// TIA Portal project "SSA-3GHz_V18" (V18) (continued)
       "SLI_gDB_T_CONFIG_PLC".configData.deviceIP.InterfaceAddress.ADDR[1] := 192;
       "SLI_gDB_T_CONFIG_PLC".configData.deviceIP.InterfaceAddress.ADDR[2] := 168;
       "SLI_gDB_T_CONFIG_PLC".configData.deviceIP.InterfaceAddress.ADDR[3] := 1;
       "SLI_gDB_T_CONFIG_PLC".configData.deviceIP.InterfaceAddress.ADDR[4] := 234;
       "SLI_gDB_T_CONFIG_PLC".configData.deviceIP.SubnetMask.ADDR[1] := 255;
       "SLI_gDB_T_CONFIG_PLC".configData.deviceIP.SubnetMask.ADDR[2] := 255;
       "SLI_gDB_T_CONFIG_PLC".configData.deviceIP.SubnetMask.ADDR[3] := 255;
       "SLI_gDB_T_CONFIG_PLC".configData.deviceIP.SubnetMask.ADDR[4] := 0;
       "SLI_gDB_T_CONFIG_PLC".configData.deviceIP.DefaultRouter.ADDR[1] := 192;
       "SLI_gDB_T_CONFIG_PLC".configData.deviceIP.DefaultRouter.ADDR[2] := 168;
       "SLI_gDB_T_CONFIG_PLC".configData.deviceIP.DefaultRouter.ADDR[3] := 1;
       "SLI_gDB_T_CONFIG_PLC".configData.deviceIP.DefaultRouter.ADDR[4] := 1;
   END_IF;
END_REGION

REGION Network 2: Set "start" to TRUE to configure the PROFINET interface.
   #_w1 := "tmp_setIP" AND NOT "Pulse_mem";   // rising edge of "tmp_setIP"
   "Pulse_mem" := "tmp_setIP";
   #_w2 := #_w1 OR "Set_IP_PArameters" OR "FirstScan" OR "RestoreFactorySettings";
   IF #_w2 THEN
       "SLI_gDB_T_CONFIG_PLC".T_CONFIG.start := TRUE;
       "Set_IP_PArameters" := FALSE;
   END_IF;
   "IEC_Timer_0_DB".TP(IN := #_w2, PT := t#5s);
   "ModbusData".serverData.disconnect := "IEC_Timer_0_DB".Q;
END_REGION

REGION Network 3: Set "start" to TRUE to configure the PROFINET interface.
   // NOTE! Before using the example:
   // 
   // Condition:
   // 1) Open the device view of the CPU "> Properties > PROFINET interface > Ethernet addresses > PROFINET". 
   // 2) To set the device name: Activate the following options: 
   // - "IP address is set directly at the device". 
   // - "PROFINET device name is set directly at the device".
   // 
   // Regarding parameter INTERFACE ("hwid"):
   // - Change the value of "hwid" according to the identification number of the PROFINET interface of your local device (CPU). (Open "PLC tags > Show all tags > System constants. Look for a name like "<Local~PROFINET_interface_1>" with a Data type "Hw_Interface". The cell "value" contains the hwid.)
   // 
   // Info:
   // In the "header" (IF_CONF_HEADER):
   // - SubfieldCount = 2: Indicates that two additional structures ("deviceIP" and "deviceName") are used below.
   // 
   // In the structure "deviceIP" (system data type IF_CONF_v4):
   // - Lenght = 18: Information on overall length of the structure (12 bytes for the device IP + 6 bytes for the parameters Id, Length and Mode)
   // - Mode = 1: Permanent change of the device IP.
   // - InterfaceAddress, SubnetMask, DefaultRouter: IP connection data.
   // 
   // In the structure "deviceName" (system data type IF_CONF_NOS):
   // - Lenght = 11: Information on overall length of the structure (5 bytes for the device name "myplc" + 6 bytes for the parameters Id, Length and Mode)
   // - Mode = 1: Permanent change of the device name in "myplc".
   // - NOS[1] ... NOS[5]: Device name (1 character / byte)
   // 
   // Note: Instead of an absolute length, you can use the default start value (Lenght = 0) for a dynamic length.
   // ENO of a box is taken as its EN; it also drops when the box reports an error
   "T_CONFIG_DB_PLC"(Req := "SLI_gDB_T_CONFIG_PLC".T_CONFIG.start,   // T_CONFIG
                     Interface := "SLI_gDB_T_CONFIG_PLC".T_CONFIG.hwid,
                     Conf_Data := "SLI_gDB_T_CONFIG_PLC".configData,
                     Done => #done_PLC,
                     Busy => "SLI_gDB_T_CONFIG_PLC".T_CONFIG.busy,
                     Error => "SLI_gDB_T_CONFIG_PLC".T_CONFIG.error,
                     Status => "SLI_gDB_T_CONFIG_PLC".T_CONFIG.status,
                     Err_Loc => #errorLocation_PLC);
   IF #done_PLC THEN "SLI_gDB_T_CONFIG_PLC".T_CONFIG.done := TRUE; END_IF;
END_REGION

REGION Network 4: INFO: Saves the value of "T_CONFIG.status" in case of an error of T_CONFIG in "T_CONFIG.memErrStat".
   RUNG wire#powerrail
      Contact( "SLI_gDB_T_CONFIG_PLC".T_CONFIG.error )
      Move(in := "SLI_gDB_T_CONFIG_PLC".T_CONFIG.status, out1 => "SLI_gDB_T_CONFIG_PLC".T_CONFIG.memErrStat)
      Move(in := #errorLocation_PLC, out1 => "SLI_gDB_T_CONFIG_PLC".T_CONFIG.errorLocation)
      R_Coil( "SLI_gDB_T_CONFIG_PLC".T_CONFIG.start )
   END_RUNG
   // the same network as SCL:
   IF "SLI_gDB_T_CONFIG_PLC".T_CONFIG.error THEN
       "SLI_gDB_T_CONFIG_PLC".T_CONFIG.memErrStat := "SLI_gDB_T_CONFIG_PLC".T_CONFIG.status;
       "SLI_gDB_T_CONFIG_PLC".T_CONFIG.errorLocation := #errorLocation_PLC;
       "SLI_gDB_T_CONFIG_PLC".T_CONFIG.start := FALSE;
   END_IF;
END_REGION

REGION Network 5: INFO: If T_CONFIG is done, "start" will be reset.
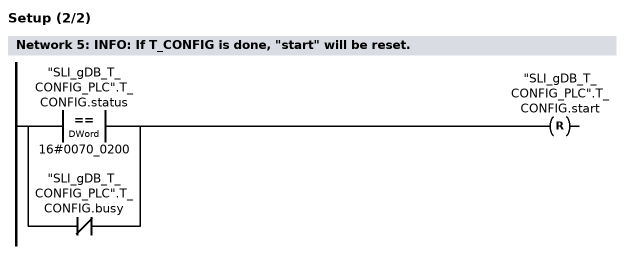
   RUNG wire#powerrail
      { S7_Templates := "SrcType := DWord" } EQ_Contact(in1 := "SLI_gDB_T_CONFIG_PLC".T_CONFIG.status, in2 := 16#0070_0200)
      wire#w1
      R_Coil( "SLI_gDB_T_CONFIG_PLC".T_CONFIG.start )
   END_RUNG
   RUNG wire#powerrail
      I_Contact( "SLI_gDB_T_CONFIG_PLC".T_CONFIG.busy )
   END_RUNG wire#w1
   // the same network as SCL:
   IF ("SLI_gDB_T_CONFIG_PLC".T_CONFIG.status = 16#0070_0200) OR NOT "SLI_gDB_T_CONFIG_PLC".T_CONFIG.busy THEN
       "SLI_gDB_T_CONFIG_PLC".T_CONFIG.start := FALSE;
   END_IF;
END_REGION
END_FUNCTION

FUNCTION "ProcessDI" : Void   // FC400, LAD
{ S7_Optimized_Access := 'TRUE' }
VERSION : 0.1
BEGIN

REGION Network 1: DutyCycOK
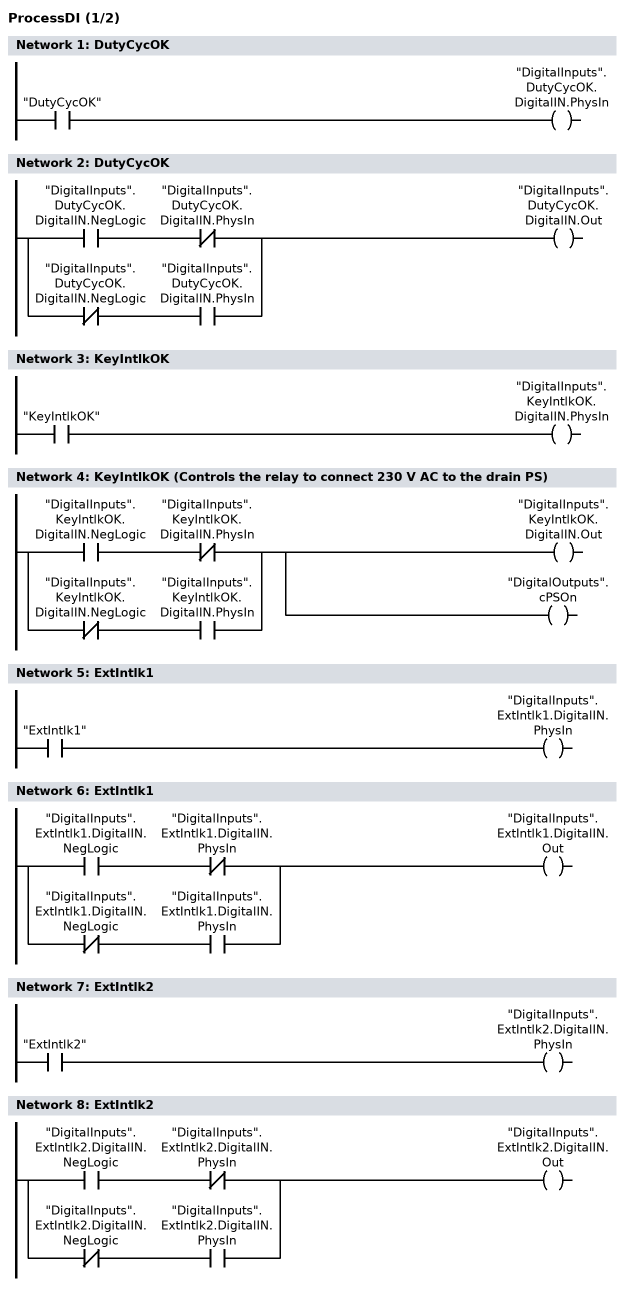
   RUNG wire#powerrail
      Contact( "DutyCycOK" )
      Coil( "DigitalInputs".DutyCycOK.DigitalIN.PhysIn )
   END_RUNG
   // the same network as SCL:
   "DigitalInputs".DutyCycOK.DigitalIN.PhysIn := "DutyCycOK";
END_REGION

REGION Network 2: DutyCycOK
   RUNG wire#powerrail
      Contact( "DigitalInputs".DutyCycOK.DigitalIN.NegLogic )
      I_Contact( "DigitalInputs".DutyCycOK.DigitalIN.PhysIn )
      wire#w1
      Coil( "DigitalInputs".DutyCycOK.DigitalIN.Out )
   END_RUNG
   RUNG wire#powerrail
      I_Contact( "DigitalInputs".DutyCycOK.DigitalIN.NegLogic )
      Contact( "DigitalInputs".DutyCycOK.DigitalIN.PhysIn )
   END_RUNG wire#w1
   // the same network as SCL:
   "DigitalInputs".DutyCycOK.DigitalIN.Out := ("DigitalInputs".DutyCycOK.DigitalIN.NegLogic AND NOT "DigitalInputs".DutyCycOK.DigitalIN.PhysIn) OR (NOT "DigitalInputs".DutyCycOK.DigitalIN.NegLogic AND "DigitalInputs".DutyCycOK.DigitalIN.PhysIn);
END_REGION

REGION Network 3: KeyIntlkOK
   RUNG wire#powerrail
      Contact( "KeyIntlkOK" )
      Coil( "DigitalInputs".KeyIntlkOK.DigitalIN.PhysIn )
   END_RUNG
   // the same network as SCL:
   "DigitalInputs".KeyIntlkOK.DigitalIN.PhysIn := "KeyIntlkOK";
END_REGION

REGION Network 4: KeyIntlkOK (Controls the relay to connect 230 V AC to the drain PS)
   RUNG wire#powerrail
      Contact( "DigitalInputs".KeyIntlkOK.DigitalIN.NegLogic )
      I_Contact( "DigitalInputs".KeyIntlkOK.DigitalIN.PhysIn )
      wire#w1
      Coil( "DigitalInputs".KeyIntlkOK.DigitalIN.Out )
   END_RUNG
   RUNG wire#powerrail
      I_Contact( "DigitalInputs".KeyIntlkOK.DigitalIN.NegLogic )
      Contact( "DigitalInputs".KeyIntlkOK.DigitalIN.PhysIn )
   END_RUNG wire#w1
   RUNG wire#w1
      Coil( "DigitalOutputs".cPSOn )
   END_RUNG
   // the same network as SCL:
   "DigitalInputs".KeyIntlkOK.DigitalIN.Out := ("DigitalInputs".KeyIntlkOK.DigitalIN.NegLogic AND NOT "DigitalInputs".KeyIntlkOK.DigitalIN.PhysIn) OR (NOT "DigitalInputs".KeyIntlkOK.DigitalIN.NegLogic AND "DigitalInputs".KeyIntlkOK.DigitalIN.PhysIn);
   "DigitalOutputs".cPSOn := "DigitalInputs".KeyIntlkOK.DigitalIN.Out;
END_REGION

REGION Network 5: ExtIntlk1
   RUNG wire#powerrail
      Contact( "ExtIntlk1" )
      Coil( "DigitalInputs".ExtIntlk1.DigitalIN.PhysIn )
   END_RUNG
   // the same network as SCL:
   "DigitalInputs".ExtIntlk1.DigitalIN.PhysIn := "ExtIntlk1";
END_REGION

REGION Network 6: ExtIntlk1
   RUNG wire#powerrail
      Contact( "DigitalInputs".ExtIntlk1.DigitalIN.NegLogic )
      I_Contact( "DigitalInputs".ExtIntlk1.DigitalIN.PhysIn )
      wire#w1
      Coil( "DigitalInputs".ExtIntlk1.DigitalIN.Out )
   END_RUNG
   RUNG wire#powerrail
      I_Contact( "DigitalInputs".ExtIntlk1.DigitalIN.NegLogic )
      Contact( "DigitalInputs".ExtIntlk1.DigitalIN.PhysIn )
   END_RUNG wire#w1
   // the same network as SCL:
   "DigitalInputs".ExtIntlk1.DigitalIN.Out := ("DigitalInputs".ExtIntlk1.DigitalIN.NegLogic AND NOT "DigitalInputs".ExtIntlk1.DigitalIN.PhysIn) OR (NOT "DigitalInputs".ExtIntlk1.DigitalIN.NegLogic AND "DigitalInputs".ExtIntlk1.DigitalIN.PhysIn);
END_REGION

REGION Network 7: ExtIntlk2
   RUNG wire#powerrail
      Contact( "ExtIntlk2" )
      Coil( "DigitalInputs".ExtIntlk2.DigitalIN.PhysIn )
   END_RUNG
   // the same network as SCL:
   "DigitalInputs".ExtIntlk2.DigitalIN.PhysIn := "ExtIntlk2";
END_REGION

REGION Network 8: ExtIntlk2
   RUNG wire#powerrail
      Contact( "DigitalInputs".ExtIntlk2.DigitalIN.NegLogic )
      I_Contact( "DigitalInputs".ExtIntlk2.DigitalIN.PhysIn )
      wire#w1
      Coil( "DigitalInputs".ExtIntlk2.DigitalIN.Out )
   END_RUNG
   RUNG wire#powerrail
      I_Contact( "DigitalInputs".ExtIntlk2.DigitalIN.NegLogic )
      Contact( "DigitalInputs".ExtIntlk2.DigitalIN.PhysIn )
   END_RUNG wire#w1
   // the same network as SCL:
   "DigitalInputs".ExtIntlk2.DigitalIN.Out := ("DigitalInputs".ExtIntlk2.DigitalIN.NegLogic AND NOT "DigitalInputs".ExtIntlk2.DigitalIN.PhysIn) OR (NOT "DigitalInputs".ExtIntlk2.DigitalIN.NegLogic AND "DigitalInputs".ExtIntlk2.DigitalIN.PhysIn);
END_REGION

REGION Network 9: T1_OK
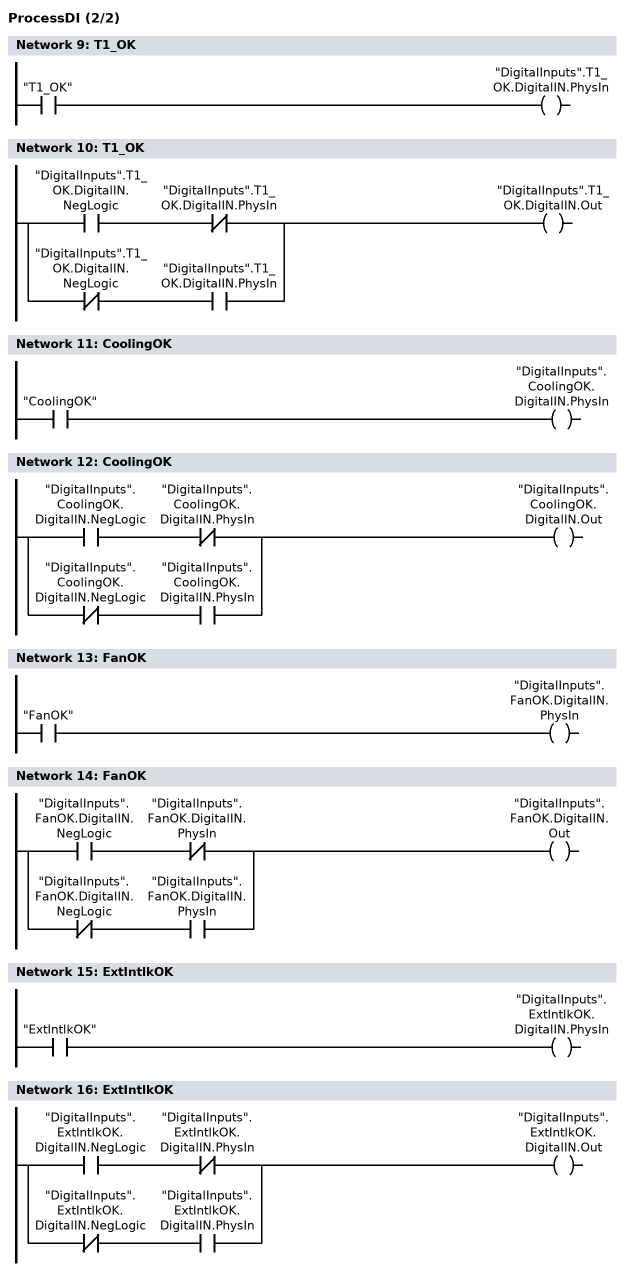
   RUNG wire#powerrail
      Contact( "T1_OK" )
      Coil( "DigitalInputs".T1_OK.DigitalIN.PhysIn )
   END_RUNG
   // the same network as SCL:
   "DigitalInputs".T1_OK.DigitalIN.PhysIn := "T1_OK";
END_REGION

REGION Network 10: T1_OK
   RUNG wire#powerrail
      Contact( "DigitalInputs".T1_OK.DigitalIN.NegLogic )
      I_Contact( "DigitalInputs".T1_OK.DigitalIN.PhysIn )
      wire#w1
      Coil( "DigitalInputs".T1_OK.DigitalIN.Out )
   END_RUNG
   RUNG wire#powerrail
      I_Contact( "DigitalInputs".T1_OK.DigitalIN.NegLogic )
      Contact( "DigitalInputs".T1_OK.DigitalIN.PhysIn )
   END_RUNG wire#w1
   // the same network as SCL:
   "DigitalInputs".T1_OK.DigitalIN.Out := ("DigitalInputs".T1_OK.DigitalIN.NegLogic AND NOT "DigitalInputs".T1_OK.DigitalIN.PhysIn) OR (NOT "DigitalInputs".T1_OK.DigitalIN.NegLogic AND "DigitalInputs".T1_OK.DigitalIN.PhysIn);
END_REGION

REGION Network 11: CoolingOK
   RUNG wire#powerrail
      Contact( "CoolingOK" )
      Coil( "DigitalInputs".CoolingOK.DigitalIN.PhysIn )
   END_RUNG
   // the same network as SCL:
   "DigitalInputs".CoolingOK.DigitalIN.PhysIn := "CoolingOK";
END_REGION

REGION Network 12: CoolingOK
   RUNG wire#powerrail
      Contact( "DigitalInputs".CoolingOK.DigitalIN.NegLogic )
      I_Contact( "DigitalInputs".CoolingOK.DigitalIN.PhysIn )
      wire#w1
      Coil( "DigitalInputs".CoolingOK.DigitalIN.Out )
   END_RUNG
   RUNG wire#powerrail
      I_Contact( "DigitalInputs".CoolingOK.DigitalIN.NegLogic )
      Contact( "DigitalInputs".CoolingOK.DigitalIN.PhysIn )
   END_RUNG wire#w1
   // the same network as SCL:
   "DigitalInputs".CoolingOK.DigitalIN.Out := ("DigitalInputs".CoolingOK.DigitalIN.NegLogic AND NOT "DigitalInputs".CoolingOK.DigitalIN.PhysIn) OR (NOT "DigitalInputs".CoolingOK.DigitalIN.NegLogic AND "DigitalInputs".CoolingOK.DigitalIN.PhysIn);
END_REGION

REGION Network 13: FanOK
   RUNG wire#powerrail
      Contact( "FanOK" )
      Coil( "DigitalInputs".FanOK.DigitalIN.PhysIn )
   END_RUNG
   // the same network as SCL:
   "DigitalInputs".FanOK.DigitalIN.PhysIn := "FanOK";
END_REGION

REGION Network 14: FanOK
   RUNG wire#powerrail
      Contact( "DigitalInputs".FanOK.DigitalIN.NegLogic )
      I_Contact( "DigitalInputs".FanOK.DigitalIN.PhysIn )
      wire#w1
      Coil( "DigitalInputs".FanOK.DigitalIN.Out )
   END_RUNG
   RUNG wire#powerrail
      I_Contact( "DigitalInputs".FanOK.DigitalIN.NegLogic )
      Contact( "DigitalInputs".FanOK.DigitalIN.PhysIn )
   END_RUNG wire#w1
   // the same network as SCL:
   "DigitalInputs".FanOK.DigitalIN.Out := ("DigitalInputs".FanOK.DigitalIN.NegLogic AND NOT "DigitalInputs".FanOK.DigitalIN.PhysIn) OR (NOT "DigitalInputs".FanOK.DigitalIN.NegLogic AND "DigitalInputs".FanOK.DigitalIN.PhysIn);
END_REGION

REGION Network 15: ExtIntlkOK
   RUNG wire#powerrail
      Contact( "ExtIntlkOK" )
      Coil( "DigitalInputs".ExtIntlkOK.DigitalIN.PhysIn )
   END_RUNG
   // the same network as SCL:
   "DigitalInputs".ExtIntlkOK.DigitalIN.PhysIn := "ExtIntlkOK";
END_REGION

REGION Network 16: ExtIntlkOK
   RUNG wire#powerrail
      Contact( "DigitalInputs".ExtIntlkOK.DigitalIN.NegLogic )
      I_Contact( "DigitalInputs".ExtIntlkOK.DigitalIN.PhysIn )
      wire#w1
      Coil( "DigitalInputs".ExtIntlkOK.DigitalIN.Out )
   END_RUNG
   RUNG wire#powerrail
      I_Contact( "DigitalInputs".ExtIntlkOK.DigitalIN.NegLogic )
      Contact( "DigitalInputs".ExtIntlkOK.DigitalIN.PhysIn )
   END_RUNG wire#w1
   // the same network as SCL:
   "DigitalInputs".ExtIntlkOK.DigitalIN.Out := ("DigitalInputs".ExtIntlkOK.DigitalIN.NegLogic AND NOT "DigitalInputs".ExtIntlkOK.DigitalIN.PhysIn) OR (NOT "DigitalInputs".ExtIntlkOK.DigitalIN.NegLogic AND "DigitalInputs".ExtIntlkOK.DigitalIN.PhysIn);
END_REGION
END_FUNCTION

FUNCTION "ProcessAI" : Void   // FC401, LAD
{ S7_Optimized_Access := 'TRUE' }
VERSION : 0.1
   VAR_TEMP
      tmpR1 : Real;
      tmpR : Real;
   END_VAR
BEGIN

REGION Network 1: U drain_RBK
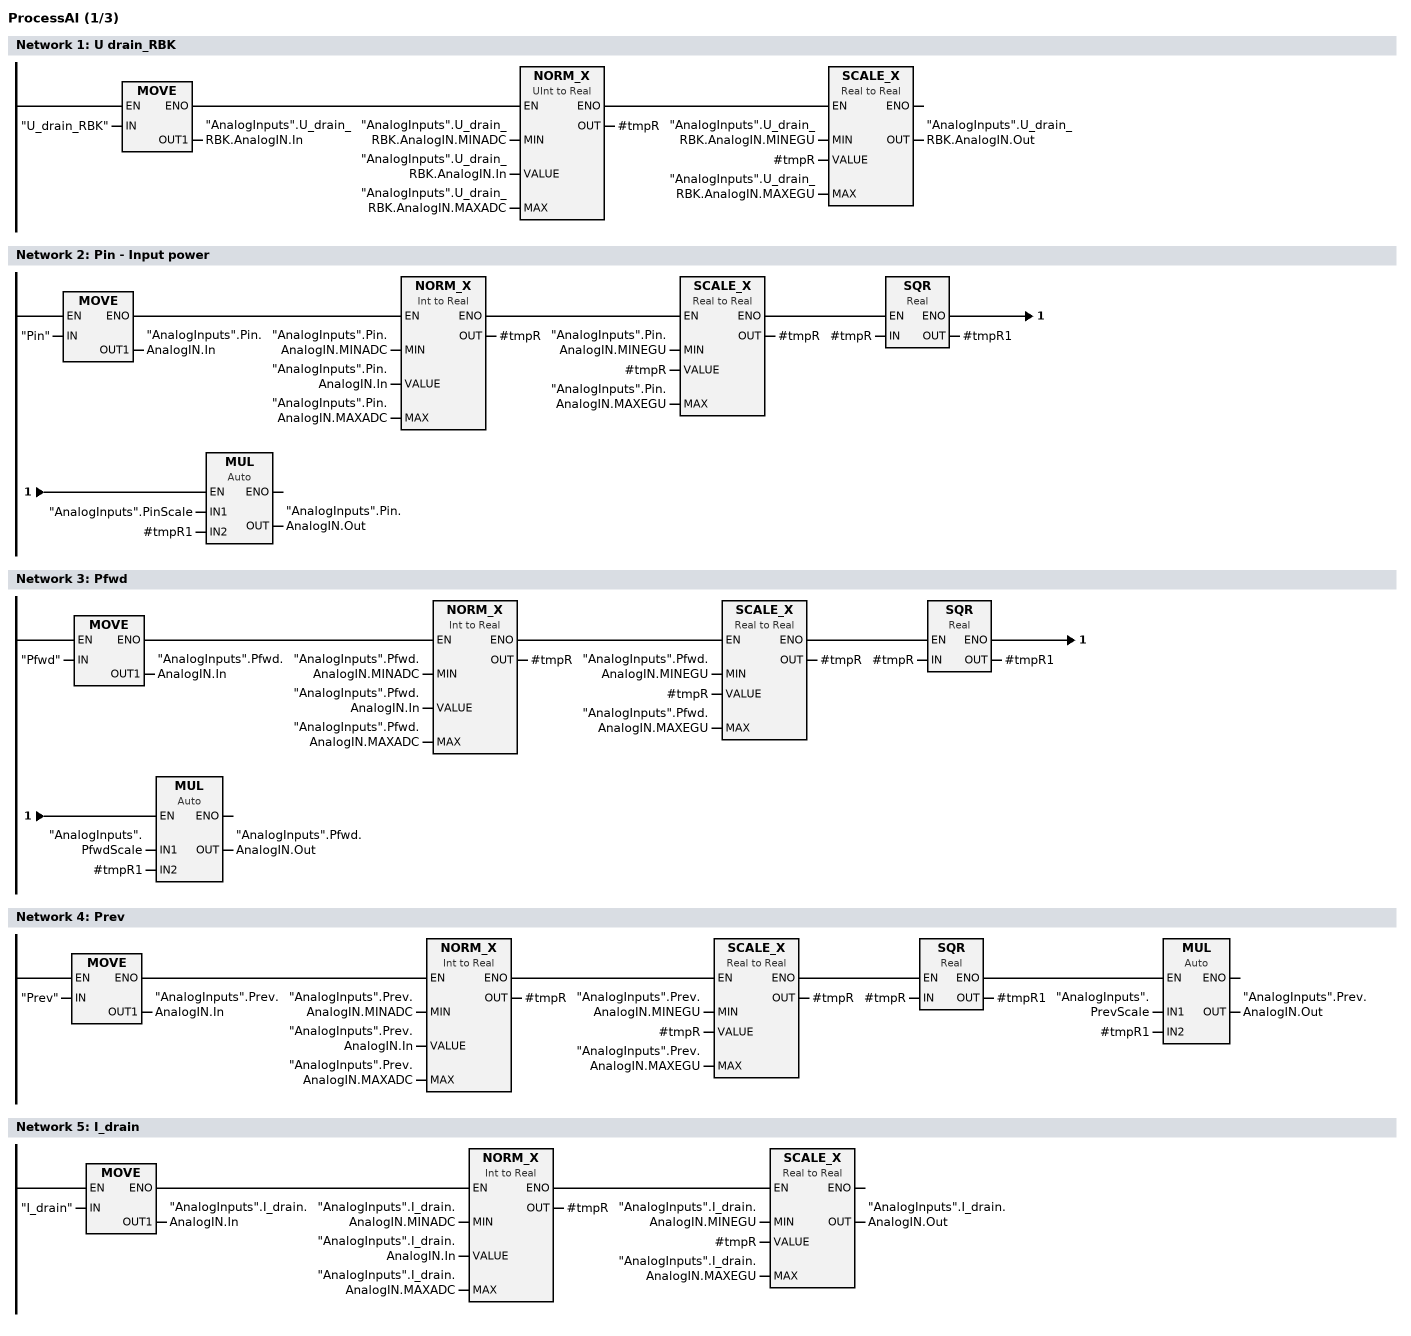
   RUNG wire#powerrail
      Move(in := "U_drain_RBK", out1 => "AnalogInputs".U_drain_RBK.AnalogIN.In)
      { S7_Templates := "[SrcType := UInt, DestType := Real]" } Normalize(min := "AnalogInputs".U_drain_RBK.AnalogIN.MINADC, value := "AnalogInputs".U_drain_RBK.AnalogIN.In, max := "AnalogInputs".U_drain_RBK.AnalogIN.MAXADC, out => #tmpR)
      { S7_Templates := "[SrcType := Real, DestType := Real]" } Scale(min := "AnalogInputs".U_drain_RBK.AnalogIN.MINEGU, value := #tmpR, max := "AnalogInputs".U_drain_RBK.AnalogIN.MAXEGU, out => "AnalogInputs".U_drain_RBK.AnalogIN.Out)
   END_RUNG
   // the same network as SCL:
   "AnalogInputs".U_drain_RBK.AnalogIN.In := "U_drain_RBK";
   #tmpR := NORM_X(MIN := "AnalogInputs".U_drain_RBK.AnalogIN.MINADC, VALUE := "AnalogInputs".U_drain_RBK.AnalogIN.In, MAX := "AnalogInputs".U_drain_RBK.AnalogIN.MAXADC);
   "AnalogInputs".U_drain_RBK.AnalogIN.Out := SCALE_X(MIN := "AnalogInputs".U_drain_RBK.AnalogIN.MINEGU, VALUE := #tmpR, MAX := "AnalogInputs".U_drain_RBK.AnalogIN.MAXEGU);
END_REGION

REGION Network 2: Pin - Input power
   "AnalogInputs".Pin.AnalogIN.In := "Pin";
   #tmpR := NORM_X(MIN := "AnalogInputs".Pin.AnalogIN.MINADC, VALUE := "AnalogInputs".Pin.AnalogIN.In, MAX := "AnalogInputs".Pin.AnalogIN.MAXADC);
   #tmpR := SCALE_X(MIN := "AnalogInputs".Pin.AnalogIN.MINEGU, VALUE := #tmpR, MAX := "AnalogInputs".Pin.AnalogIN.MAXEGU);
   #tmpR1 := SQR(#tmpR);
   "AnalogInputs".Pin.AnalogIN.Out := "AnalogInputs".PinScale * #tmpR1;
END_REGION

REGION Network 3: Pfwd
   "AnalogInputs".Pfwd.AnalogIN.In := "Pfwd";
   #tmpR := NORM_X(MIN := "AnalogInputs".Pfwd.AnalogIN.MINADC, VALUE := "AnalogInputs".Pfwd.AnalogIN.In, MAX := "AnalogInputs".Pfwd.AnalogIN.MAXADC);
   #tmpR := SCALE_X(MIN := "AnalogInputs".Pfwd.AnalogIN.MINEGU, VALUE := #tmpR, MAX := "AnalogInputs".Pfwd.AnalogIN.MAXEGU);
   #tmpR1 := SQR(#tmpR);
   "AnalogInputs".Pfwd.AnalogIN.Out := "AnalogInputs".PfwdScale * #tmpR1;
END_REGION

REGION Network 4: Prev
   "AnalogInputs".Prev.AnalogIN.In := "Prev";
   #tmpR := NORM_X(MIN := "AnalogInputs".Prev.AnalogIN.MINADC, VALUE := "AnalogInputs".Prev.AnalogIN.In, MAX := "AnalogInputs".Prev.AnalogIN.MAXADC);
   #tmpR := SCALE_X(MIN := "AnalogInputs".Prev.AnalogIN.MINEGU, VALUE := #tmpR, MAX := "AnalogInputs".Prev.AnalogIN.MAXEGU);
   #tmpR1 := SQR(#tmpR);
   "AnalogInputs".Prev.AnalogIN.Out := "AnalogInputs".PrevScale * #tmpR1;
END_REGION

REGION Network 5: I_drain
   RUNG wire#powerrail
      Move(in := "I_drain", out1 => "AnalogInputs".I_drain.AnalogIN.In)
      { S7_Templates := "[SrcType := Int, DestType := Real]" } Normalize(min := "AnalogInputs".I_drain.AnalogIN.MINADC, value := "AnalogInputs".I_drain.AnalogIN.In, max := "AnalogInputs".I_drain.AnalogIN.MAXADC, out => #tmpR)
      { S7_Templates := "[SrcType := Real, DestType := Real]" } Scale(min := "AnalogInputs".I_drain.AnalogIN.MINEGU, value := #tmpR, max := "AnalogInputs".I_drain.AnalogIN.MAXEGU, out => "AnalogInputs".I_drain.AnalogIN.Out)
   END_RUNG
   // the same network as SCL:
   "AnalogInputs".I_drain.AnalogIN.In := "I_drain";
   #tmpR := NORM_X(MIN := "AnalogInputs".I_drain.AnalogIN.MINADC, VALUE := "AnalogInputs".I_drain.AnalogIN.In, MAX := "AnalogInputs".I_drain.AnalogIN.MAXADC);
   "AnalogInputs".I_drain.AnalogIN.Out := SCALE_X(MIN := "AnalogInputs".I_drain.AnalogIN.MINEGU, VALUE := #tmpR, MAX := "AnalogInputs".I_drain.AnalogIN.MAXEGU);
END_REGION

REGION Network 6: ADC0ch1
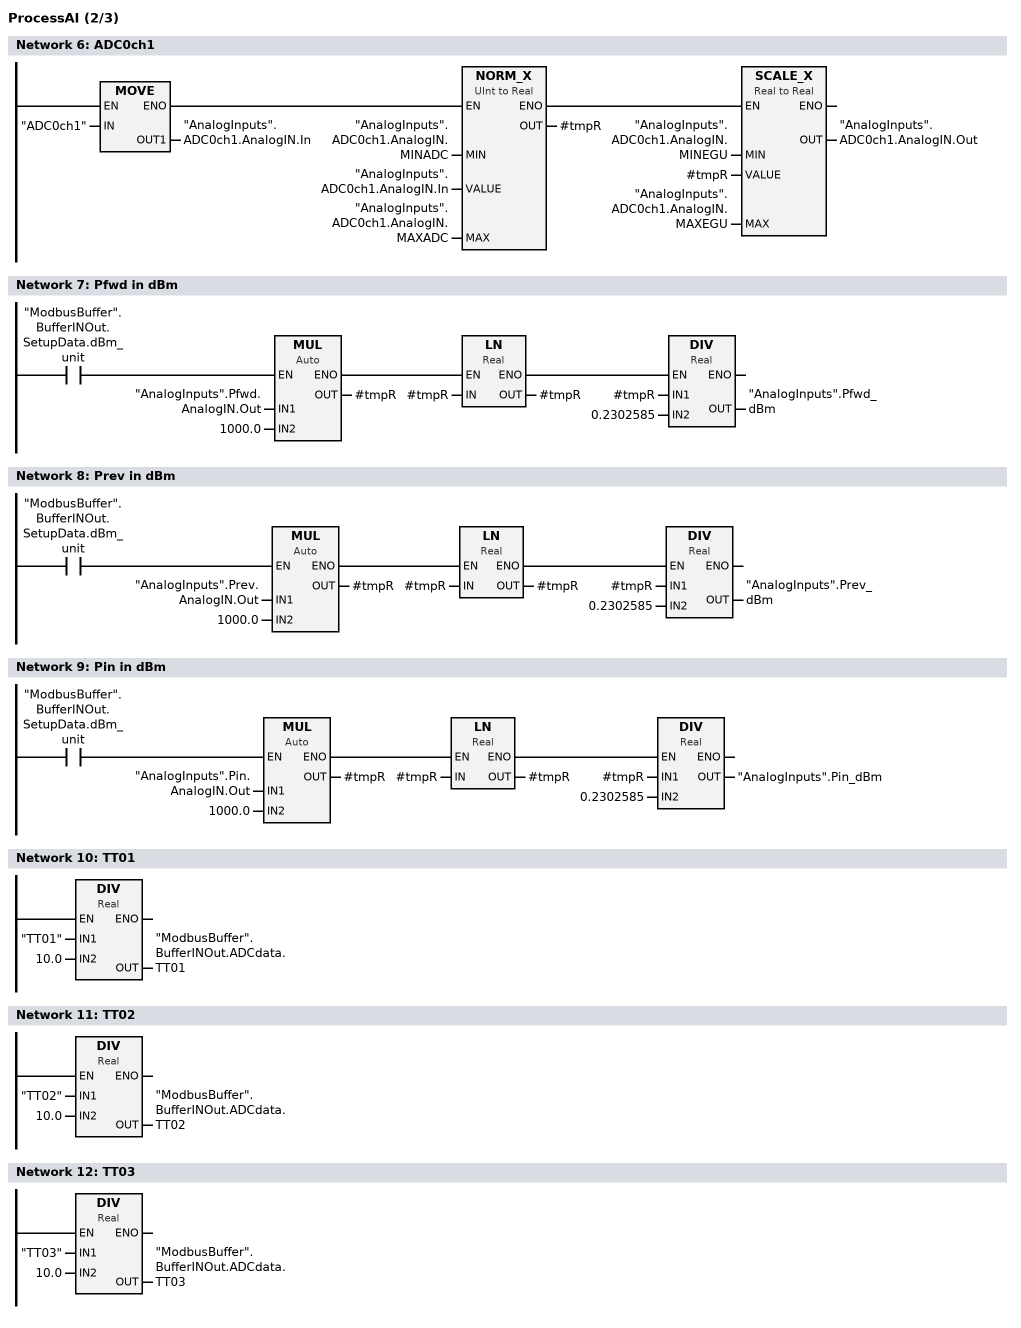
   RUNG wire#powerrail
      Move(in := "ADC0ch1", out1 => "AnalogInputs".ADC0ch1.AnalogIN.In)
      { S7_Templates := "[SrcType := UInt, DestType := Real]" } Normalize(min := "AnalogInputs".ADC0ch1.AnalogIN.MINADC, value := "AnalogInputs".ADC0ch1.AnalogIN.In, max := "AnalogInputs".ADC0ch1.AnalogIN.MAXADC, out => #tmpR)
      { S7_Templates := "[SrcType := Real, DestType := Real]" } Scale(min := "AnalogInputs".ADC0ch1.AnalogIN.MINEGU, value := #tmpR, max := "AnalogInputs".ADC0ch1.AnalogIN.MAXEGU, out => "AnalogInputs".ADC0ch1.AnalogIN.Out)
   END_RUNG
   // the same network as SCL:
   "AnalogInputs".ADC0ch1.AnalogIN.In := "ADC0ch1";
   #tmpR := NORM_X(MIN := "AnalogInputs".ADC0ch1.AnalogIN.MINADC, VALUE := "AnalogInputs".ADC0ch1.AnalogIN.In, MAX := "AnalogInputs".ADC0ch1.AnalogIN.MAXADC);
   "AnalogInputs".ADC0ch1.AnalogIN.Out := SCALE_X(MIN := "AnalogInputs".ADC0ch1.AnalogIN.MINEGU, VALUE := #tmpR, MAX := "AnalogInputs".ADC0ch1.AnalogIN.MAXEGU);
END_REGION

REGION Network 7: Pfwd in dBm
   IF "ModbusBuffer".BufferINOut.SetupData.dBm_unit THEN
       #tmpR := "AnalogInputs".Pfwd.AnalogIN.Out * 1000.0;
       #tmpR := LN(#tmpR);
       "AnalogInputs".Pfwd_dBm := #tmpR / 0.2302585;
   END_IF;
END_REGION

REGION Network 8: Prev in dBm
   IF "ModbusBuffer".BufferINOut.SetupData.dBm_unit THEN
       #tmpR := "AnalogInputs".Prev.AnalogIN.Out * 1000.0;
       #tmpR := LN(#tmpR);
       "AnalogInputs".Prev_dBm := #tmpR / 0.2302585;
   END_IF;
END_REGION

REGION Network 9: Pin in dBm
   IF "ModbusBuffer".BufferINOut.SetupData.dBm_unit THEN
       #tmpR := "AnalogInputs".Pin.AnalogIN.Out * 1000.0;
       #tmpR := LN(#tmpR);
       "AnalogInputs".Pin_dBm := #tmpR / 0.2302585;
   END_IF;
END_REGION

REGION Network 10: TT01
   RUNG wire#powerrail
      { S7_Templates := "SrcType := Real" } Div(in1 := "TT01", in2 := 10.0, out => "ModbusBuffer".BufferINOut.ADCdata.TT01)
   END_RUNG
   // the same network as SCL:
   "ModbusBuffer".BufferINOut.ADCdata.TT01 := "TT01" / 10.0;
END_REGION

REGION Network 11: TT02
   RUNG wire#powerrail
      { S7_Templates := "SrcType := Real" } Div(in1 := "TT02", in2 := 10.0, out => "ModbusBuffer".BufferINOut.ADCdata.TT02)
   END_RUNG
   // the same network as SCL:
   "ModbusBuffer".BufferINOut.ADCdata.TT02 := "TT02" / 10.0;
END_REGION

REGION Network 12: TT03
   RUNG wire#powerrail
      { S7_Templates := "SrcType := Real" } Div(in1 := "TT03", in2 := 10.0, out => "ModbusBuffer".BufferINOut.ADCdata.TT03)
   END_RUNG
   // the same network as SCL:
   "ModbusBuffer".BufferINOut.ADCdata.TT03 := "TT03" / 10.0;
END_REGION

REGION Network 13: TT04
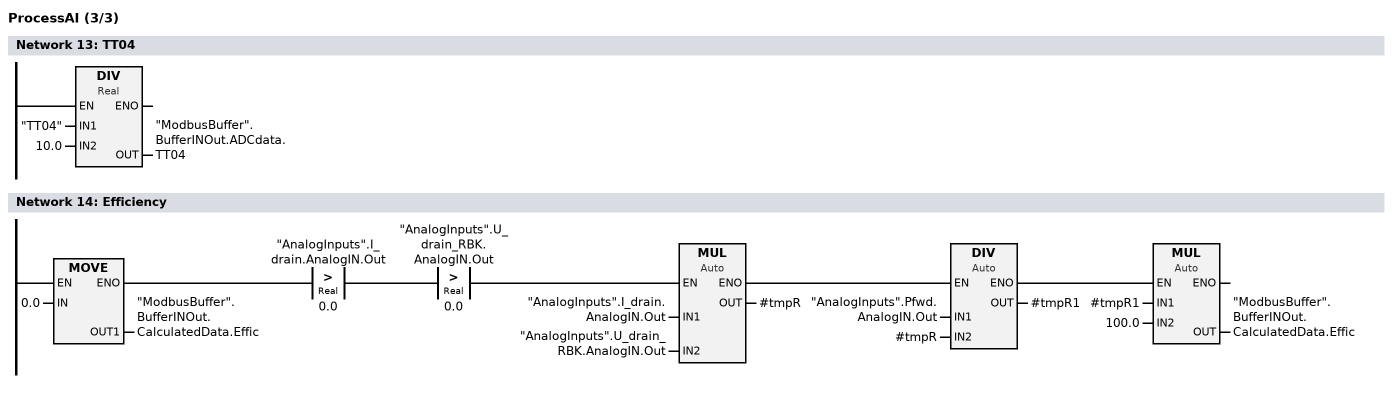
   RUNG wire#powerrail
      { S7_Templates := "SrcType := Real" } Div(in1 := "TT04", in2 := 10.0, out => "ModbusBuffer".BufferINOut.ADCdata.TT04)
   END_RUNG
   // the same network as SCL:
   "ModbusBuffer".BufferINOut.ADCdata.TT04 := "TT04" / 10.0;
END_REGION

REGION Network 14: Efficiency
   RUNG wire#powerrail
      Move(in := 0.0, out1 => "ModbusBuffer".BufferINOut.CalculatedData.Effic)
      { S7_Templates := "SrcType := Real" } GT_Contact(in1 := "AnalogInputs".I_drain.AnalogIN.Out, in2 := 0.0)
      { S7_Templates := "SrcType := Real" } GT_Contact(in1 := "AnalogInputs".U_drain_RBK.AnalogIN.Out, in2 := 0.0)
      Mul(in1 := "AnalogInputs".I_drain.AnalogIN.Out, in2 := "AnalogInputs".U_drain_RBK.AnalogIN.Out, out => #tmpR)
      Div(in1 := "AnalogInputs".Pfwd.AnalogIN.Out, in2 := #tmpR, out => #tmpR1)
      Mul(in1 := #tmpR1, in2 := 100.0, out => "ModbusBuffer".BufferINOut.CalculatedData.Effic)
   END_RUNG
   // the same network as SCL:
   "ModbusBuffer".BufferINOut.CalculatedData.Effic := 0.0;
   IF ("AnalogInputs".I_drain.AnalogIN.Out > 0.0) AND ("AnalogInputs".U_drain_RBK.AnalogIN.Out > 0.0) THEN
       #tmpR := "AnalogInputs".I_drain.AnalogIN.Out * "AnalogInputs".U_drain_RBK.AnalogIN.Out;
       #tmpR1 := "AnalogInputs".Pfwd.AnalogIN.Out / #tmpR;
       "ModbusBuffer".BufferINOut.CalculatedData.Effic := #tmpR1 * 100.0;
   END_IF;
END_REGION
END_FUNCTION

FUNCTION "ProcessAO" : Void   // FC402, LAD
{ S7_Optimized_Access := 'TRUE' }
VERSION : 0.1
   VAR_TEMP
      tmpR : Real;
   END_VAR
BEGIN

REGION Network 1: U drain
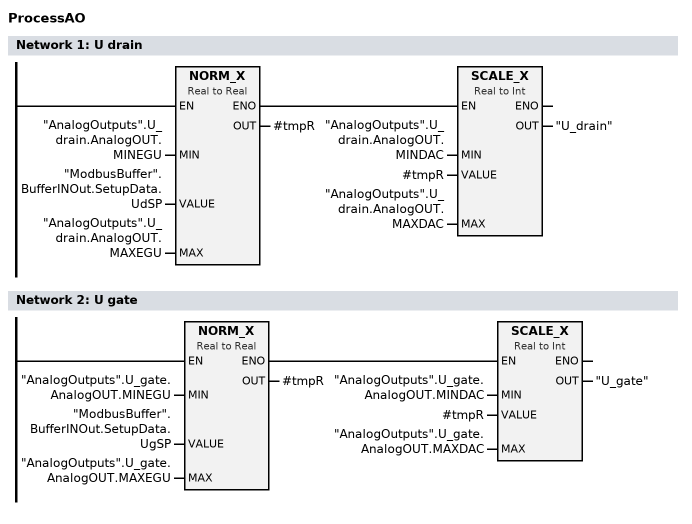
   RUNG wire#powerrail
      { S7_Templates := "[SrcType := Real, DestType := Real]" } Normalize(min := "AnalogOutputs".U_drain.AnalogOUT.MINEGU, value := "ModbusBuffer".BufferINOut.SetupData.UdSP, max := "AnalogOutputs".U_drain.AnalogOUT.MAXEGU, out => #tmpR)
      { S7_Templates := "[SrcType := Real, DestType := Int]" } Scale(min := "AnalogOutputs".U_drain.AnalogOUT.MINDAC, value := #tmpR, max := "AnalogOutputs".U_drain.AnalogOUT.MAXDAC, out => "U_drain")
   END_RUNG
   // the same network as SCL:
   #tmpR := NORM_X(MIN := "AnalogOutputs".U_drain.AnalogOUT.MINEGU, VALUE := "ModbusBuffer".BufferINOut.SetupData.UdSP, MAX := "AnalogOutputs".U_drain.AnalogOUT.MAXEGU);
   "U_drain" := SCALE_X(MIN := "AnalogOutputs".U_drain.AnalogOUT.MINDAC, VALUE := #tmpR, MAX := "AnalogOutputs".U_drain.AnalogOUT.MAXDAC);
END_REGION

REGION Network 2: U gate
   RUNG wire#powerrail
      { S7_Templates := "[SrcType := Real, DestType := Real]" } Normalize(min := "AnalogOutputs".U_gate.AnalogOUT.MINEGU, value := "ModbusBuffer".BufferINOut.SetupData.UgSP, max := "AnalogOutputs".U_gate.AnalogOUT.MAXEGU, out => #tmpR)
      { S7_Templates := "[SrcType := Real, DestType := Int]" } Scale(min := "AnalogOutputs".U_gate.AnalogOUT.MINDAC, value := #tmpR, max := "AnalogOutputs".U_gate.AnalogOUT.MAXDAC, out => "U_gate")
   END_RUNG
   // the same network as SCL:
   #tmpR := NORM_X(MIN := "AnalogOutputs".U_gate.AnalogOUT.MINEGU, VALUE := "ModbusBuffer".BufferINOut.SetupData.UgSP, MAX := "AnalogOutputs".U_gate.AnalogOUT.MAXEGU);
   "U_gate" := SCALE_X(MIN := "AnalogOutputs".U_gate.AnalogOUT.MINDAC, VALUE := #tmpR, MAX := "AnalogOutputs".U_gate.AnalogOUT.MAXDAC);
END_REGION
END_FUNCTION

FUNCTION "ProcessDO" : Void   // FC450, LAD
{ S7_Optimized_Access := 'TRUE' }
VERSION : 0.1
BEGIN

REGION Network 1: RF switcch
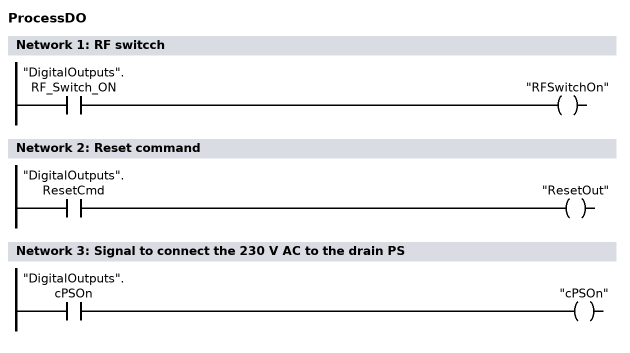
   RUNG wire#powerrail
      Contact( "DigitalOutputs".RF_Switch_ON )
      Coil( "RFSwitchOn" )
   END_RUNG
   // the same network as SCL:
   "RFSwitchOn" := "DigitalOutputs".RF_Switch_ON;
END_REGION

REGION Network 2: Reset command
   RUNG wire#powerrail
      Contact( "DigitalOutputs".ResetCmd )
      Coil( "ResetOut" )
   END_RUNG
   // the same network as SCL:
   "ResetOut" := "DigitalOutputs".ResetCmd;
END_REGION

REGION Network 3: Signal to connect the 230 V AC to the drain PS
   RUNG wire#powerrail
      Contact( "DigitalOutputs".cPSOn )
      Coil( "cPSOn" )
   END_RUNG
   // the same network as SCL:
   "cPSOn" := "DigitalOutputs".cPSOn;
END_REGION
END_FUNCTION

FUNCTION "CalcTransistorV" : Void   // FC500, SCL
{ S7_Optimized_Access := 'TRUE' }
VERSION : 0.1
   VAR_INPUT
      NominalPwr : Real;
      size : Int;   // max size if the lookup table. Valid data until Pwr != 0
   END_VAR
   VAR_OUTPUT
      UdSP : Real;
      UgSP : Real;
   END_VAR
   VAR_TEMP
      Pwr : Real;
      Ud : Real;
      Ug : Real;
      K : Real;
      i : Int;
   END_VAR
BEGIN
   (*
   Calculate the Darin and gate voltages based on the nominal power
   *)
   IF "ModbusBuffer".BufferINOut.SetupData.dBm_unit THEN
       "ModbusBuffer".BufferINOut.SetupData.NominalPower := EXP("ModbusBuffer".BufferINOut.SetupData.NominalPower_dBm* 0.2302585) / 1000.0;
   ELSE
       "ModbusBuffer".BufferINOut.SetupData.NominalPower_dBm := 10.0 * LN(1000.0 *"ModbusBuffer".BufferINOut.SetupData.NominalPower)/ 2.302585;
   END_IF;

   IF #NominalPwr <= "ModbusBuffer".BufferINOut.LookupTable.Pwr[0] THEN
       #UdSP := "ModbusBuffer".BufferINOut.LookupTable.Ud[0];
       #UgSP := "ModbusBuffer".BufferINOut.LookupTable.Ug[0];
   ELSE
       FOR #i := 1 TO #size-1 DO
       // Statement section FOR
           #Pwr := "ModbusBuffer".BufferINOut.LookupTable.Pwr[#i];
           IF #Pwr = 0 THEN
               //the end of table marker
               #UdSP := "ModbusBuffer".BufferINOut.LookupTable.Ud[#i - 1];
               #UgSP := "ModbusBuffer".BufferINOut.LookupTable.Ug[#i - 1];
               RETURN;
           END_IF;
           IF #NominalPwr > #Pwr THEN
               CONTINUE;
           END_IF;
           #K := (#NominalPwr - "ModbusBuffer".BufferINOut.LookupTable.Pwr[#i - 1]) / (#Pwr - "ModbusBuffer".BufferINOut.LookupTable.Pwr[#i - 1]);
           #UdSP := "ModbusBuffer".BufferINOut.LookupTable.Ud[#i-1] + #K * ("ModbusBuffer".BufferINOut.LookupTable.Ud[#i] - "ModbusBuffer".BufferINOut.LookupTable.Ud[#i-1]);
           #UgSP := "ModbusBuffer".BufferINOut.LookupTable.Ug[#i - 1] + #K * ("ModbusBuffer".BufferINOut.LookupTable.Ug[#i] - "ModbusBuffer".BufferINOut.LookupTable.Ug[#i - 1]);
           RETURN;
       END_FOR;
       #UdSP := "ModbusBuffer".BufferINOut.LookupTable.Ud[#size-1];
       #UgSP := "ModbusBuffer".BufferINOut.LookupTable.Ug[#size-1];
   END_IF;
END_FUNCTION

FUNCTION "Interlocks" : Void   // FC600, LAD
{ S7_Optimized_Access := 'TRUE' }
VERSION : 0.1
BEGIN

REGION Network 1: RF Switch